         CALL  "#FC_CONTROL_HEATER"
         ( TtA      := "IOC2PLC".TT600,
           TtB      := "IOC2PLC".TT670,
           TtC      := "IOC2PLC".TT680,
           TtD      := "IOC2PLC".TT690,
           TtE      := #Unused_TT,
           TtF      := #Unused_TT,
           Nb_Tt    := 4,
           TS       := #TS,
           ExtCmd   := #ExtCmd,
           cmdEpics := "Epics_to_PLC"."EH60_67-69",
           EH       := "voie 5 chaufferette BV",
           sEpics   := "PLC_to_Epics"."EH60_67-69",
           Object   := "#DATA_HEATERS"."EH60_67-69"
         );
END_REGION

REGION Network 7 (STL): EH97-98 - VB channel 6
   // Dewar, Electrical Heater
         L     2;
         T     "#DATA_HEATERS"."EH97-98".P_TS_Ton;
         T     "#DATA_HEATERS"."EH97-98".P_Pilot_Ton;
         L     5;
         T     "#DATA_HEATERS"."EH97-98".P_TS_Toff;

         SET;
         A     "IOC2PLC".TT970_VALID;
         A     "IOC2PLC".TT980_VALID;
         A     "EPICS_COMM_OK";
         =     #TS;
   // Force the heater ON when the temperature data is not valid
   // (TS = FALSE). The heater will be turned on for 30 s and TS
   // will be forced TRUE for 30 s. This will hopefully raise the
   // temperature enough for Pt100 to be in range (>73 K)
         SET;
         AN    #TS;
         A(;
         A     "#DATA_HEATERS"."EH97-98".XH;
         A     "#DATA_HEATERS"."EH97-98".X;
         O;
         AN    "#DATA_HEATERS"."EH97-98".XH;
         A     "#DATA_HEATERS"."EH97-98".H;
         );
         =     #ExtCmdTrig;
         CALL  TP , "IEC_Timer_EH97-98_DB"
         ( IN := #ExtCmdTrig,
           PT := T#30s,
           Q  := #ExtCmd,
           ET := #tmp_et
         );
         A     #ExtCmd;
         S     #TS;

         CALL  "#FC_CONTROL_HEATER"
         ( TtA      := "IOC2PLC".TT970,
           TtB      := "IOC2PLC".TT980,
           TtC      := #Unused_TT,
           TtD      := #Unused_TT,
           TtE      := #Unused_TT,
           TtF      := #Unused_TT,
           Nb_Tt    := 2,
           TS       := #TS,
           ExtCmd   := #ExtCmd,
           cmdEpics := "Epics_to_PLC"."EH97-98",
           EH       := "voie 6 chaufferette BV",
           sEpics   := "PLC_to_Epics"."EH97-98",
           Object   := "#DATA_HEATERS"."EH97-98"
         );
END_REGION

REGION Network 8 (STL): EH01 - CM channel 1
         L     2;
         T     "#DATA_HEATERS".EH01.P_TS_Ton;
         T     "#DATA_HEATERS".EH01.P_Pilot_Ton;
         L     5;
         T     "#DATA_HEATERS".EH01.P_TS_Toff;

         SET;
         A     "IOC2PLC".TT04_VALID;
         A     "IOC2PLC".TT06_VALID;
         A     "EPICS_COMM_OK";
         =     #TS;

         CALL  "#FC_CONTROL_HEATER"
         ( TtA      := "IOC2PLC".TT04,
           TtB      := "IOC2PLC".TT06,
           TtC      := #Unused_TT,
           TtD      := #Unused_TT,
           TtE      := #Unused_TT,
           TtF      := #Unused_TT,
           Nb_Tt    := 2,
           TS       := #TS,
           ExtCmd   := #ExtCmd,
           cmdEpics := "Epics_to_PLC".EH01,
           EH       := "voie 1 chaufferette CM",
           sEpics   := "PLC_to_Epics".EH01,
           Object   := "#DATA_HEATERS".EH01
         );
END_REGION

REGION Network 9 (STL): EH02 - CM channel 2
         L     2;
         T     "#DATA_HEATERS".EH02.P_TS_Ton;
         T     "#DATA_HEATERS".EH02.P_Pilot_Ton;
         L     5;
         T     "#DATA_HEATERS".EH02.P_TS_Toff;

         SET;
         A     "IOC2PLC".TT05_VALID;
         A     "IOC2PLC".TT07_VALID;
         A     "EPICS_COMM_OK";
         =     #TS;

         CALL  "#FC_CONTROL_HEATER"
         ( TtA      := "IOC2PLC".TT05,
           TtB      := "IOC2PLC".TT07,
           TtC      := #Unused_TT,
           TtD      := #Unused_TT,
           TtE      := #Unused_TT,
           TtF      := #Unused_TT,
           Nb_Tt    := 2,
           TS       := #TS,
           ExtCmd   := #ExtCmd,
           cmdEpics := "Epics_to_PLC".EH02,
           EH       := "voie 2 chaufferette CM",
           sEpics   := "PLC_to_Epics".EH02,
           Object   := "#DATA_HEATERS".EH02
         );
END_REGION

REGION Network 10 (STL): EH10 - CM channel 3
         L     2;
         T     "#DATA_HEATERS".EH10.P_TS_Ton;
         T     "#DATA_HEATERS".EH10.P_Pilot_Ton;
         L     5;
         T     "#DATA_HEATERS".EH10.P_TS_Toff;

         SET;
         A     "IOC2PLC"."CTS:TT10_VALID";
         A     "IOC2PLC"."CTS:TT11_VALID";
         A     "EPICS_COMM_OK";
         =     #TS;

         CALL  "#FC_CONTROL_HEATER"
         ( TtA      := "IOC2PLC"."CTS:TT10",
           TtB      := "IOC2PLC"."CTS:TT11",
           TtC      := #Unused_TT,
           TtD      := #Unused_TT,
           TtE      := #Unused_TT,
           TtF      := #Unused_TT,
           Nb_Tt    := 2,
           TS       := #TS,
           ExtCmd   := #ExtCmd,
           cmdEpics := "Epics_to_PLC".EH10,
           EH       := "voie 3 chaufferette CM",
           sEpics   := "PLC_to_Epics".EH10,
           Object   := "#DATA_HEATERS".EH10
         );
END_REGION

REGION Network 11 (STL): EH20 - CM channel 4
         L     2;
         T     "#DATA_HEATERS".EH20.P_TS_Ton;
         T     "#DATA_HEATERS".EH20.P_Pilot_Ton;
         L     5;
         T     "#DATA_HEATERS".EH20.P_TS_Toff;

         SET;
         A     "IOC2PLC"."CTS:TT20_VALID";
         A     "IOC2PLC"."CTS:TT21_VALID";
         A     "EPICS_COMM_OK";
         =     #TS;

         CALL  "#FC_CONTROL_HEATER"
         ( TtA      := "IOC2PLC"."CTS:TT20",
           TtB      := "IOC2PLC"."CTS:TT21",
           TtC      := #Unused_TT,
           TtD      := #Unused_TT,
           TtE      := #Unused_TT,
           TtF      := #Unused_TT,
           Nb_Tt    := 2,
           TS       := #TS,
           ExtCmd   := #ExtCmd,
           cmdEpics := "Epics_to_PLC".EH20,
           EH       := "voie 4 chaufferette CM",
           sEpics   := "PLC_to_Epics".EH20,
           Object   := "#DATA_HEATERS".EH20
         );
END_REGION

REGION Network 12 (STL): EH918 - CM channel 9
   // Dewar, Electrical Heater
         L     2;
         T     "#DATA_HEATERS"."spare-CM-9".P_TS_Ton;
         T     "#DATA_HEATERS"."spare-CM-9".P_Pilot_Ton;
         L     5;
         T     "#DATA_HEATERS"."spare-CM-9".P_TS_Toff;

         SET;
         A     "IOC2PLC"."CTS:TT20_VALID";
         A     "EPICS_COMM_OK";
         =     #TS;
   // Force the heater ON when the temperature data is not valid
   // (TS = FALSE). The heater will be turned on for 30 s and TS
   // will be forced TRUE for 30 s. This will hopefully raise the
   // temperature enough for Pt100 to be in range (>73 K)
         SET;
         AN    #TS;
         A(;
         A     "#DATA_HEATERS"."spare-CM-9".XH;
         A     "#DATA_HEATERS"."spare-CM-9".X;
         O;
         AN    "#DATA_HEATERS"."spare-CM-9".XH;
         A     "#DATA_HEATERS"."spare-CM-9".H;
         );
         =     #ExtCmdTrig;
         CALL  TP , "IEC_Timer_EH918_DB"
         ( IN := #ExtCmdTrig,
           PT := T#30s,
           Q  := #ExtCmd,
           ET := #tmp_et
         );
         A     #ExtCmd;
         S     #TS;

   _191: CALL  "#FC_CONTROL_HEATER"
         ( TtA      := "IOC2PLC"."CTS:TT20",
           TtB      := #Unused_TT,
           TtC      := #Unused_TT,
           TtD      := #Unused_TT,
           TtE      := #Unused_TT,
           TtF      := #Unused_TT,
           Nb_Tt    := 1,
           TS       := #TS,
           ExtCmd   := #ExtCmd,
           cmdEpics := "Epics_to_PLC"."spare-CM-9",
           EH       := "voie 9 chaufferette CM",
           sEpics   := "PLC_to_Epics"."spare-CM-9",
           Object   := "#DATA_HEATERS"."spare-CM-9"
         );
END_REGION

REGION Network 13 (STL): EH904 - CM channel 11
   // Dewar, Electrical Heater
         L     2;
         T     "#DATA_HEATERS"."spare-CM-11".P_TS_Ton;
         T     "#DATA_HEATERS"."spare-CM-11".P_Pilot_Ton;
         L     5;
         T     "#DATA_HEATERS"."spare-CM-11".P_TS_Toff;

         SET;
         A     "IOC2PLC"."CTS:TT21_VALID";
         A     "EPICS_COMM_OK";
         =     #TS;

   // Force the heater ON when the temperature data is not valid
   // (TS = FALSE). The heater will be turned on for 30 s and TS
   // will be forced TRUE for 30 s. This will hopefully raise the
   // temperature enough for Pt100 to be in range (>73 K)
         SET;
         AN    #TS;
         A(;
         A     "#DATA_HEATERS"."spare-CM-11".XH;
         A     "#DATA_HEATERS"."spare-CM-11".X;
         O;
         AN    "#DATA_HEATERS"."spare-CM-11".XH;
         A     "#DATA_HEATERS"."spare-CM-11".H;
         );
         =     #ExtCmdTrig;
         CALL  TP , "IEC_Timer_EH904_DB"
         ( IN := #ExtCmdTrig,
           PT := T#30s,
           Q  := #ExtCmd,
           ET := #tmp_et
         );
         A     #ExtCmd;
         S     #TS;

         CALL  "#FC_CONTROL_HEATER"
         ( TtA      := "IOC2PLC"."CTS:TT21",
           TtB      := #Unused_TT,
           TtC      := #Unused_TT,
           TtD      := #Unused_TT,
           TtE      := #Unused_TT,
           TtF      := #Unused_TT,
           Nb_Tt    := 1,
           TS       := #TS,
           ExtCmd   := #ExtCmd,
           cmdEpics := "Epics_to_PLC"."spare-CM-11",
           EH       := "voie 11 chaufferette CM",
           sEpics   := "PLC_to_Epics"."spare-CM-11",
           Object   := "#DATA_HEATERS"."spare-CM-11"
         );
END_REGION

REGION Network 14 (STL): EH12 - Coupler 1 flange
   // Dewar, Electrical Heater
         L     2;
         T     "#DATA_HEATERS".EH12.P_TS_Ton;
         T     "#DATA_HEATERS".EH12.P_Pilot_Ton;
         L     5;
         T     "#DATA_HEATERS".EH12.P_TS_Toff;

         L     "PLC_to_Epics".TT120.Visu;
         L     0;
         ==I;
         =     #Enable;
         CALL  "#FC_CONTROL_HEATER"
         ( TtA      := "PLC_to_Epics".TT120.Level,
           TtB      := #Unused_TT,
           TtC      := #Unused_TT,
           TtD      := #Unused_TT,
           TtE      := #Unused_TT,
           TtF      := #Unused_TT,
           Nb_Tt    := 1,
           TS       := #Enable,
           ExtCmd   := #ExtCmd,
           cmdEpics := "Epics_to_PLC".EH12,
           EH       := "EH12 Cpl1",
           sEpics   := "PLC_to_Epics".EH12,
           Object   := "#DATA_HEATERS".EH12
         );
END_REGION

REGION Network 15 (STL): EH22 - Coupler 2 flange
   // Dewar, Electrical Heater
         L     2;
         T     "#DATA_HEATERS".EH22.P_TS_Ton;
         T     "#DATA_HEATERS".EH22.P_Pilot_Ton;
         L     5;
         T     "#DATA_HEATERS".EH22.P_TS_Toff;

         L     "PLC_to_Epics".TT220.Visu;
         L     0;
         ==I;
         =     #Enable;
         CALL  "#FC_CONTROL_HEATER"
         ( TtA      := "PLC_to_Epics".TT220.Level,
           TtB      := #Unused_TT,
           TtC      := #Unused_TT,
           TtD      := #Unused_TT,
           TtE      := #Unused_TT,
           TtF      := #Unused_TT,
           Nb_Tt    := 1,
           TS       := #Enable,
           ExtCmd   := #ExtCmd,
           cmdEpics := "Epics_to_PLC".EH22,
           EH       := "EH22 Cpl2",
           sEpics   := "PLC_to_Epics".EH22,
           Object   := "#DATA_HEATERS".EH22
         );
END_REGION
END_FUNCTION

FUNCTION "Manage_HEATERS" : Void   // FC513, LAD
TITLE = Manage the heaters
{ S7_Optimized_Access := 'FALSE' }
AUTHOR : KG
VERSION : 0.1
BEGIN

REGION Network 1: EH12 & EH22 - Coupler flange cavity 1 and 2
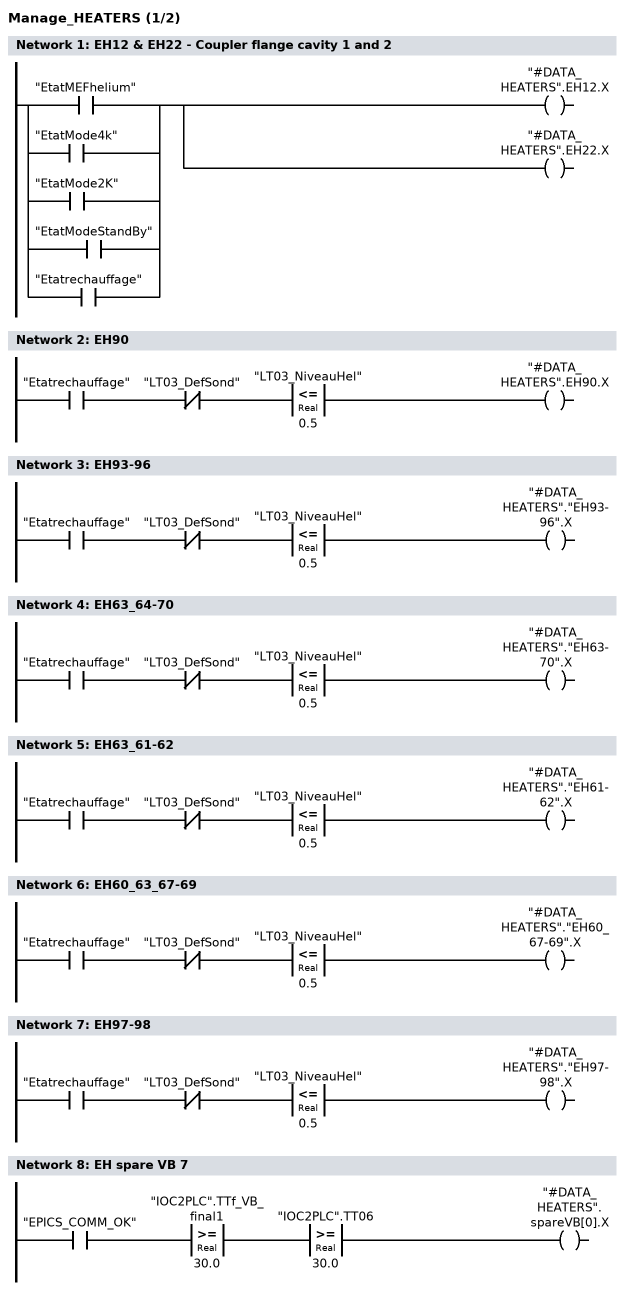
   RUNG wire#powerrail
      Contact( "EtatMEFhelium" )
      wire#w1
      Coil( "#DATA_HEATERS".EH12.X )
   END_RUNG
   RUNG wire#powerrail
      Contact( "EtatMode4k" )
   END_RUNG wire#w1
   RUNG wire#powerrail
      Contact( "EtatMode2K" )
   END_RUNG wire#w1
   RUNG wire#powerrail
      Contact( "EtatModeStandBy" )
   END_RUNG wire#w1
   RUNG wire#powerrail
      Contact( "Etatrechauffage" )
   END_RUNG wire#w1
   RUNG wire#w1
      Coil( "#DATA_HEATERS".EH22.X )
   END_RUNG
   // the same network as SCL:
   "#DATA_HEATERS".EH12.X := "EtatMEFhelium" OR "EtatMode4k" OR "EtatMode2K" OR "EtatModeStandBy" OR "Etatrechauffage";
   "#DATA_HEATERS".EH22.X := "#DATA_HEATERS".EH12.X;
END_REGION

REGION Network 2: EH90
   RUNG wire#powerrail
      Contact( "Etatrechauffage" )
      I_Contact( "LT03_DefSond" )
      { S7_Templates := "SrcType := Real" } LE_Contact(in1 := "LT03_NiveauHel", in2 := 0.5)
      Coil( "#DATA_HEATERS".EH90.X )
   END_RUNG
   // the same network as SCL:
   "#DATA_HEATERS".EH90.X := "Etatrechauffage" AND NOT "LT03_DefSond" AND ("LT03_NiveauHel" <= 0.5);
END_REGION

REGION Network 3: EH93-96
   RUNG wire#powerrail
      Contact( "Etatrechauffage" )
      I_Contact( "LT03_DefSond" )
      { S7_Templates := "SrcType := Real" } LE_Contact(in1 := "LT03_NiveauHel", in2 := 0.5)
      Coil( "#DATA_HEATERS"."EH93-96".X )
   END_RUNG
   // the same network as SCL:
   "#DATA_HEATERS"."EH93-96".X := "Etatrechauffage" AND NOT "LT03_DefSond" AND ("LT03_NiveauHel" <= 0.5);
END_REGION

REGION Network 4: EH63_64-70
   RUNG wire#powerrail
      Contact( "Etatrechauffage" )
      I_Contact( "LT03_DefSond" )
      { S7_Templates := "SrcType := Real" } LE_Contact(in1 := "LT03_NiveauHel", in2 := 0.5)
      Coil( "#DATA_HEATERS"."EH63-70".X )
   END_RUNG
   // the same network as SCL:
   "#DATA_HEATERS"."EH63-70".X := "Etatrechauffage" AND NOT "LT03_DefSond" AND ("LT03_NiveauHel" <= 0.5);
END_REGION

REGION Network 5: EH63_61-62
   RUNG wire#powerrail
      Contact( "Etatrechauffage" )
      I_Contact( "LT03_DefSond" )
      { S7_Templates := "SrcType := Real" } LE_Contact(in1 := "LT03_NiveauHel", in2 := 0.5)
      Coil( "#DATA_HEATERS"."EH61-62".X )
   END_RUNG
   // the same network as SCL:
   "#DATA_HEATERS"."EH61-62".X := "Etatrechauffage" AND NOT "LT03_DefSond" AND ("LT03_NiveauHel" <= 0.5);
END_REGION

REGION Network 6: EH60_63_67-69
   RUNG wire#powerrail
      Contact( "Etatrechauffage" )
      I_Contact( "LT03_DefSond" )
      { S7_Templates := "SrcType := Real" } LE_Contact(in1 := "LT03_NiveauHel", in2 := 0.5)
      Coil( "#DATA_HEATERS"."EH60_67-69".X )
   END_RUNG
   // the same network as SCL:
   "#DATA_HEATERS"."EH60_67-69".X := "Etatrechauffage" AND NOT "LT03_DefSond" AND ("LT03_NiveauHel" <= 0.5);
END_REGION

REGION Network 7: EH97-98
   RUNG wire#powerrail
      Contact( "Etatrechauffage" )
      I_Contact( "LT03_DefSond" )
      { S7_Templates := "SrcType := Real" } LE_Contact(in1 := "LT03_NiveauHel", in2 := 0.5)
      Coil( "#DATA_HEATERS"."EH97-98".X )
   END_RUNG
   // the same network as SCL:
   "#DATA_HEATERS"."EH97-98".X := "Etatrechauffage" AND NOT "LT03_DefSond" AND ("LT03_NiveauHel" <= 0.5);
END_REGION

REGION Network 8: EH spare VB 7
   RUNG wire#powerrail
      Contact( "EPICS_COMM_OK" )
      { S7_Templates := "SrcType := Real" } GE_Contact(in1 := "IOC2PLC".TTf_VB_final1, in2 := 30.0)
      { S7_Templates := "SrcType := Real" } GE_Contact(in1 := "IOC2PLC".TT06, in2 := 30.0)
      Coil( "#DATA_HEATERS".spareVB[0].X )
   END_RUNG
   // the same network as SCL:
   "#DATA_HEATERS".spareVB[0].X := "EPICS_COMM_OK" AND ("IOC2PLC".TTf_VB_final1 >= 30.0) AND ("IOC2PLC".TT06 >= 30.0);
END_REGION

REGION Network 9: EH spare CM 11
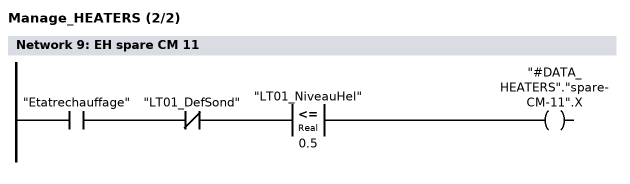
   RUNG wire#powerrail
      Contact( "Etatrechauffage" )
      I_Contact( "LT01_DefSond" )
      { S7_Templates := "SrcType := Real" } LE_Contact(in1 := "LT01_NiveauHel", in2 := 0.5)
      Coil( "#DATA_HEATERS"."spare-CM-11".X )
   END_RUNG
   // the same network as SCL:
   "#DATA_HEATERS"."spare-CM-11".X := "Etatrechauffage" AND NOT "LT01_DefSond" AND ("LT01_NiveauHel" <= 0.5);
END_REGION
END_FUNCTION

FUNCTION "Manage_VALVES" : Void   // FC556, LAD
TITLE = Manage the valves
{ S7_Optimized_Access := 'FALSE' }
AUTHOR : KG
VERSION : 0.1
BEGIN

REGION Network 1: RV90
   // Open the release valve when the pressure is over the threshold
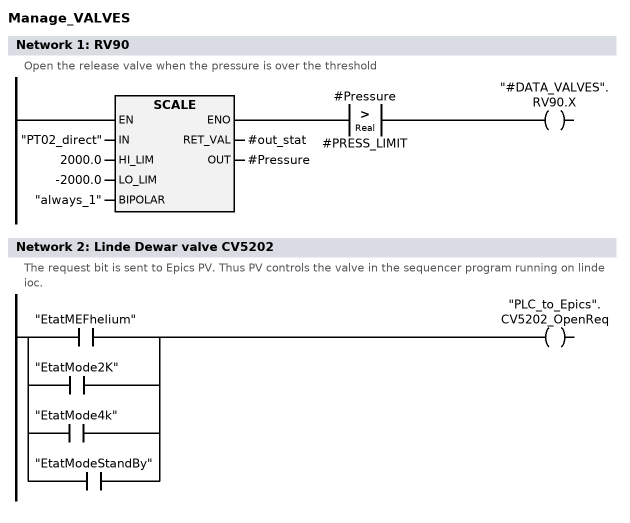
   // ENO of a box is taken as its EN; it also drops when the box reports an error
   #out_stat := SCALE(IN := "PT02_direct",
                      HI_LIM := 2000.0,
                      LO_LIM := -2000.0,
                      BIPOLAR := "always_1",
                      OUT => #Pressure);
   "#DATA_VALVES".RV90.X := #Pressure > #PRESS_LIMIT;
END_REGION

REGION Network 2: Linde Dewar valve CV5202
   // The request bit is sent to Epics PV. Thus PV controls the valve in the sequencer program running on linde ioc.
   RUNG wire#powerrail
      Contact( "EtatMEFhelium" )
      wire#w1
      Coil( "PLC_to_Epics".CV5202_OpenReq )
   END_RUNG
   RUNG wire#powerrail
      Contact( "EtatMode2K" )
   END_RUNG wire#w1
   RUNG wire#powerrail
      Contact( "EtatMode4k" )
   END_RUNG wire#w1
   RUNG wire#powerrail
      Contact( "EtatModeStandBy" )
   END_RUNG wire#w1
   // the same network as SCL:
   "PLC_to_Epics".CV5202_OpenReq := "EtatMEFhelium" OR "EtatMode2K" OR "EtatMode4k" OR "EtatModeStandBy";
END_REGION
END_FUNCTION

ORGANIZATION_BLOCK "Main"   // OB1, STL
TITLE = "Main Program Sweep (Cycle)"
{ S7_Optimized_Access := 'FALSE' }
VERSION : 0.1
BEGIN

REGION Network 1: Set-up the timing pulse for FC_TIMER
         A     "point1sec";
         AN    "point1secMem";
         =     "point1secPls";
         A     "point1sec";
         =     "point1secMem";

         SET;
         A     "oneSec";
         AN    "oneSecMem";
         =     "oneSecPls";
         A     "oneSec";
         =     "oneSecMem";
END_REGION

REGION Network 2: Get data and commands from Epics IOC
         CALL  "Recv_from_Epics";
         NOP   0;
END_REGION

REGION Network 3
         A     "Graph/manuelle";
         JNB   Label_0;
         CALL  "commande vanne";
   Label_0:NOP   0;
END_REGION

REGION Network 4
         CALL  "NIveau Helium&Pression&vide";
         NOP   0;
END_REGION

REGION Network 5
         CALL  "ACQ_CABTF";
         NOP   0;
END_REGION

REGION Network 6
         AN    "Graph/manuelle";
         JNB   Label_1;
         CALL  "grafcet";
   Label_1:NOP   0;
END_REGION

REGION Network 7
         CALL  "Send_to_Epics";
         NOP   0;
END_REGION

REGION Network 8: Instantiate the heaters control
         CALL  "INST_CONTROL_HEATER";
END_REGION

REGION Network 9: Instantiate the valve control
         CALL  "INST_VALVES";
END_REGION

REGION Network 10: Manage the heaters
         CALL  "Manage_HEATERS";
END_REGION

REGION Network 11: Manage the valves
         CALL  "Manage_VALVES";
END_REGION

REGION Network 12
         CALL  "UpdateData2HNOSS";
END_REGION

REGION Network 13: Appeler le bloc de diagnostic système / Call system diagnostics block
         CALL  "RSE_FB", "RSE_DB";
END_REGION

REGION Network 14: Clear INIT flag after the first cycle
         SET;
         R     "INIT";
END_REGION
END_ORGANIZATION_BLOCK

ORGANIZATION_BLOCK "CYC_INT2"   // OB32, LAD
TITLE = Cyclic_1s / "Cyclic Interrupt"
{ S7_Optimized_Access := 'FALSE' }
AUTHOR : KG
VERSION : 0.1
// Call the PID functionswith 1s interval
   VAR_TEMP   // added for the SCL form of the ladder/FBD networks
      _w1 : Bool;
   END_VAR
BEGIN

REGION Network 1: PID regulator for the LN2 screen cooling (CV60)
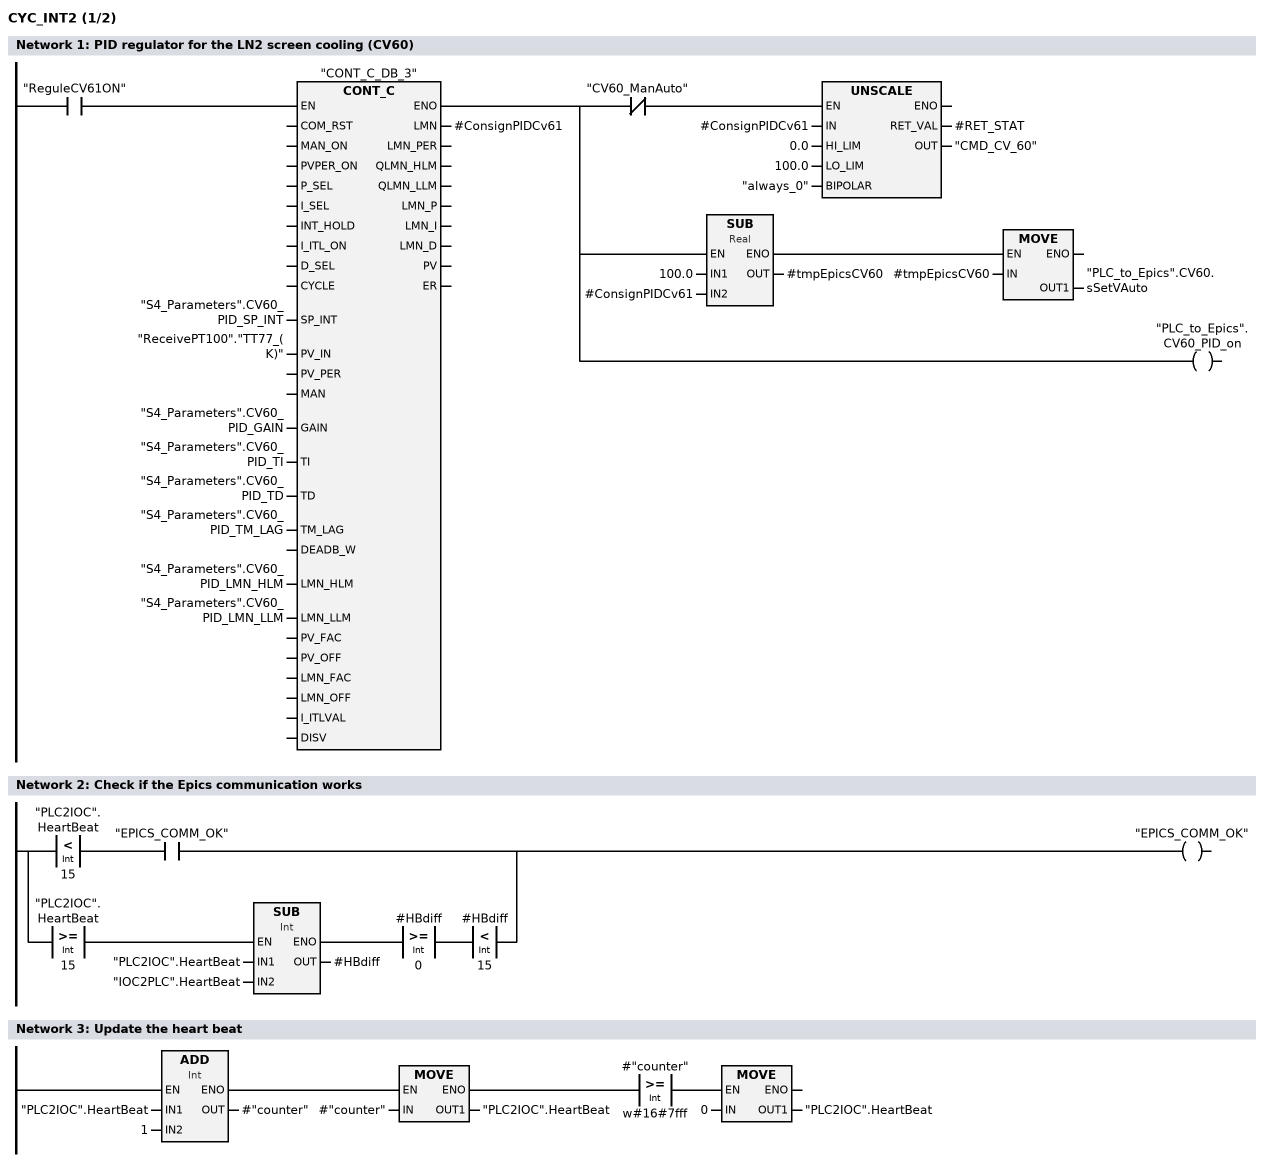
   // ENO of a box is taken as its EN; it also drops when the box reports an error
   #_w1 := "ReguleCV61ON";
   IF #_w1 THEN
       "CONT_C_DB_3"(SP_INT := "S4_Parameters".CV60_PID_SP_INT,   // CONT_C
                     PV_IN := "ReceivePT100"."TT77_(K)",
                     GAIN := "S4_Parameters".CV60_PID_GAIN,
                     TI := "S4_Parameters".CV60_PID_TI,
                     TD := "S4_Parameters".CV60_PID_TD,
                     TM_LAG := "S4_Parameters".CV60_PID_TM_LAG,
                     LMN_HLM := "S4_Parameters".CV60_PID_LMN_HLM,
                     LMN_LLM := "S4_Parameters".CV60_PID_LMN_LLM,
                     LMN => #ConsignPIDCv61);
   END_IF;
   IF #_w1 AND NOT "CV60_ManAuto" THEN
       #RET_STAT := UNSCALE(IN := #ConsignPIDCv61,
                            HI_LIM := 0.0,
                            LO_LIM := 100.0,
                            BIPOLAR := "always_0",
                            OUT => "CMD_CV_60");
   END_IF;
   IF #_w1 THEN
       #tmpEpicsCV60 := 100.0 - #ConsignPIDCv61;
       "PLC_to_Epics".CV60.sSetVAuto := #tmpEpicsCV60;
   END_IF;
   "PLC_to_Epics".CV60_PID_on := #_w1;
END_REGION

REGION Network 2: Check if the Epics communication works
   // ENO of a box is taken as its EN; it also drops when the box reports an error
   #_w1 := "PLC2IOC".HeartBeat >= 15;
   IF #_w1 THEN #HBdiff := "PLC2IOC".HeartBeat - "IOC2PLC".HeartBeat; END_IF;
   "EPICS_COMM_OK" := (#_w1 AND (#HBdiff >= 0) AND (#HBdiff < 15)) OR (("PLC2IOC".HeartBeat < 15) AND "EPICS_COMM_OK");
END_REGION

REGION Network 3: Update the heart beat
   RUNG wire#powerrail
      { S7_Templates := "SrcType := Int"; S7_GenerateENO := "TRUE" } Add(in1 := "PLC2IOC".HeartBeat, in2 := 1, out => #"counter")
      { S7_GenerateENO := "TRUE" } Move(in := #"counter", out1 => "PLC2IOC".HeartBeat)
      { S7_Templates := "SrcType := Int" } GE_Contact(in1 := #"counter", in2 := w#16#7fff)
      { S7_GenerateENO := "TRUE" } Move(in := 0, out1 => "PLC2IOC".HeartBeat)
   END_RUNG
   // the same network as SCL:
   // ENO of a box is taken as its EN; it also drops when the box reports an error
   #"counter" := "PLC2IOC".HeartBeat + 1;
   "PLC2IOC".HeartBeat := #"counter";
   IF #"counter" >= w#16#7fff THEN "PLC2IOC".HeartBeat := 0; END_IF;
END_REGION

REGION Network 4: Check if the communicationto HNOSS PLC works
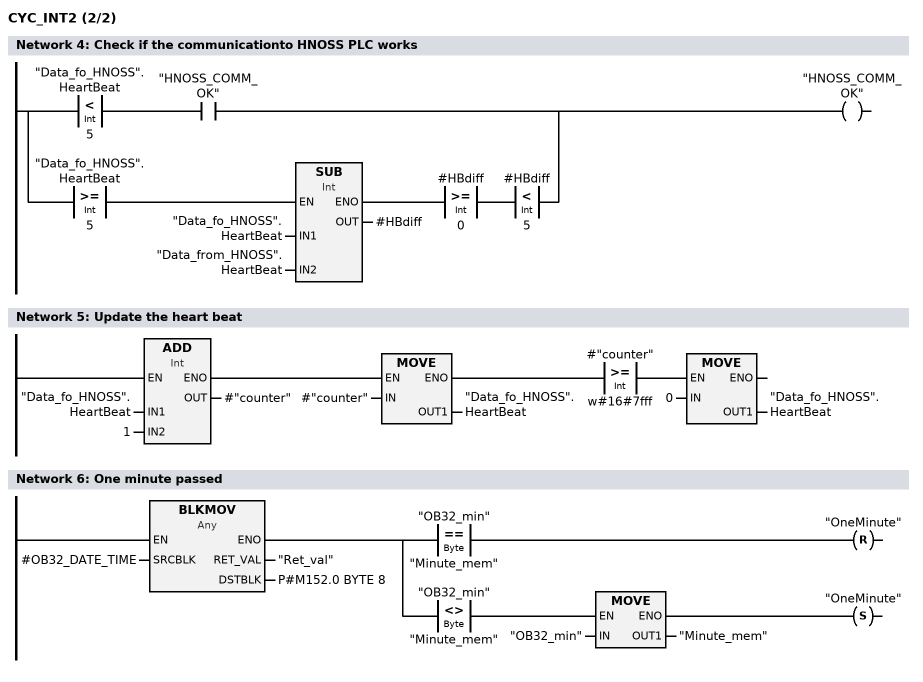
   // ENO of a box is taken as its EN; it also drops when the box reports an error
   #_w1 := "Data_fo_HNOSS".HeartBeat >= 5;
   IF #_w1 THEN #HBdiff := "Data_fo_HNOSS".HeartBeat - "Data_from_HNOSS".HeartBeat; END_IF;
   "HNOSS_COMM_OK" := (#_w1 AND (#HBdiff >= 0) AND (#HBdiff < 5)) OR (("Data_fo_HNOSS".HeartBeat < 5) AND "HNOSS_COMM_OK");
END_REGION

REGION Network 5: Update the heart beat
   RUNG wire#powerrail
      { S7_Templates := "SrcType := Int"; S7_GenerateENO := "TRUE" } Add(in1 := "Data_fo_HNOSS".HeartBeat, in2 := 1, out => #"counter")
      { S7_GenerateENO := "TRUE" } Move(in := #"counter", out1 => "Data_fo_HNOSS".HeartBeat)
      { S7_Templates := "SrcType := Int" } GE_Contact(in1 := #"counter", in2 := w#16#7fff)
      { S7_GenerateENO := "TRUE" } Move(in := 0, out1 => "Data_fo_HNOSS".HeartBeat)
   END_RUNG
   // the same network as SCL:
   // ENO of a box is taken as its EN; it also drops when the box reports an error
   #"counter" := "Data_fo_HNOSS".HeartBeat + 1;
   "Data_fo_HNOSS".HeartBeat := #"counter";
   IF #"counter" >= w#16#7fff THEN "Data_fo_HNOSS".HeartBeat := 0; END_IF;
END_REGION

REGION Network 6: One minute passed
   // ENO of a box is taken as its EN; it also drops when the box reports an error
   "Ret_val" := BLKMOV(SRCBLK := #OB32_DATE_TIME, DSTBLK => P#M152.0 BYTE 8);
   IF "OB32_min" = "Minute_mem" THEN "OneMinute" := FALSE; END_IF;
   #_w1 := "OB32_min" <> "Minute_mem";
   IF #_w1 THEN
       "Minute_mem" := "OB32_min";
       "OneMinute" := TRUE;
   END_IF;
END_REGION
END_ORGANIZATION_BLOCK

ORGANIZATION_BLOCK "CYC_INT5"   // OB35, LAD
TITLE = "Cyclic Interrupt"
{ S7_Optimized_Access := 'FALSE' }
VERSION : 0.1
// Period 100 ms
   VAR_TEMP   // added for the SCL form of the ladder/FBD networks
      _w1 : Bool;
      _w2 : Bool;
   END_VAR
BEGIN

REGION Network 1
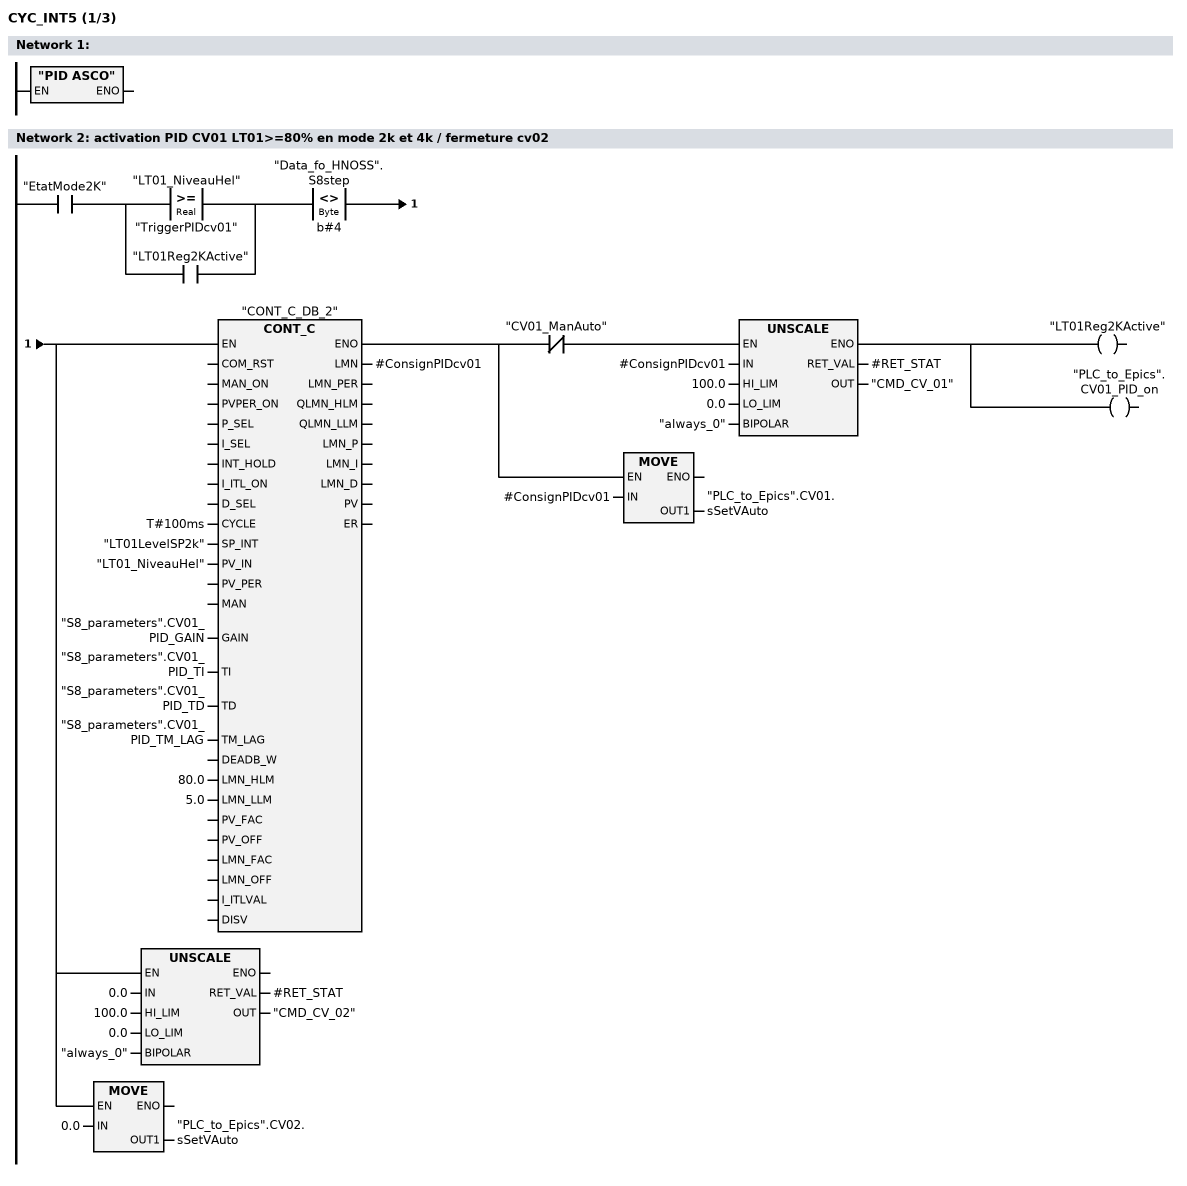
   RUNG wire#powerrail
      "PID ASCO"()
   END_RUNG
   // the same network as SCL:
   "PID ASCO"();
END_REGION

REGION Network 2: activation PID CV01 LT01>=80% en mode 2k et 4k / fermeture cv02
   // ENO of a box is taken as its EN; it also drops when the box reports an error
   #_w1 := "EtatMode2K" AND (("LT01_NiveauHel" >= "TriggerPIDcv01") OR "LT01Reg2KActive") AND ("Data_fo_HNOSS".S8step <> b#4);
   IF #_w1 THEN
       "CONT_C_DB_2"(CYCLE := T#100ms,   // CONT_C
                     SP_INT := "LT01LevelSP2k",
                     PV_IN := "LT01_NiveauHel",
                     GAIN := "S8_parameters".CV01_PID_GAIN,
                     TI := "S8_parameters".CV01_PID_TI,
                     TD := "S8_parameters".CV01_PID_TD,
                     TM_LAG := "S8_parameters".CV01_PID_TM_LAG,
                     LMN_HLM := 80.0,
                     LMN_LLM := 5.0,
                     LMN => #ConsignPIDcv01);
   END_IF;
   #_w2 := #_w1 AND NOT "CV01_ManAuto";
   IF #_w2 THEN
       #RET_STAT := UNSCALE(IN := #ConsignPIDcv01,
                            HI_LIM := 100.0,
                            LO_LIM := 0.0,
                            BIPOLAR := "always_0",
                            OUT => "CMD_CV_01");
   END_IF;
   "LT01Reg2KActive" := #_w2;
   "PLC_to_Epics".CV01_PID_on := #_w2;
   IF #_w1 THEN
       "PLC_to_Epics".CV01.sSetVAuto := #ConsignPIDcv01;
       #RET_STAT := UNSCALE(IN := 0.0, HI_LIM := 100.0, LO_LIM := 0.0, BIPOLAR := "always_0", OUT => "CMD_CV_02");
       "PLC_to_Epics".CV02.sSetVAuto := 0.0;
   END_IF;
END_REGION

REGION Network 3: activation PID CV03 LT03>=80%
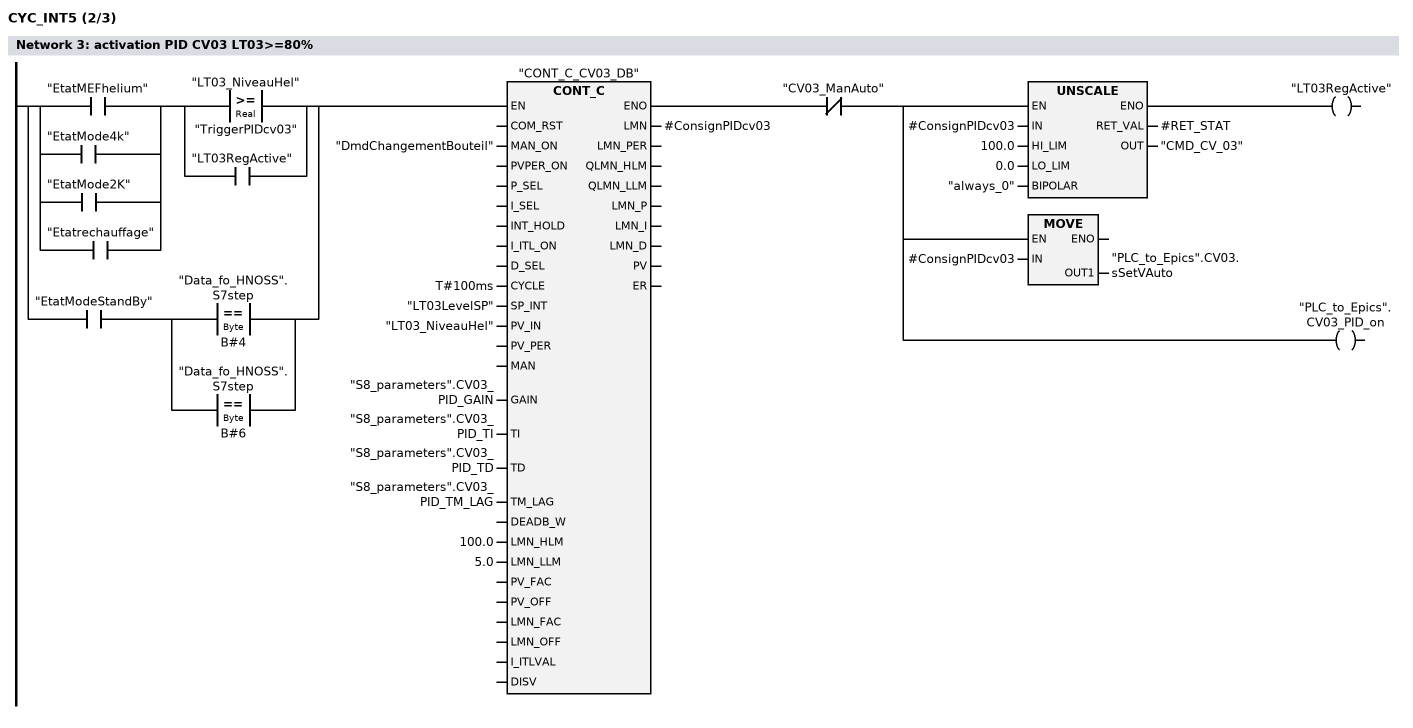
   // ENO of a box is taken as its EN; it also drops when the box reports an error
   #_w1 := (("EtatMEFhelium" OR "EtatMode4k" OR "EtatMode2K" OR "Etatrechauffage") AND (("LT03_NiveauHel" >= "TriggerPIDcv03") OR "LT03RegActive")) OR ("EtatModeStandBy" AND (("Data_fo_HNOSS".S7step = B#4) OR ("Data_fo_HNOSS".S7step = B#6)));
   IF #_w1 THEN
       "CONT_C_CV03_DB"(MAN_ON := "DmdChangementBouteil",   // CONT_C
                        CYCLE := T#100ms,
                        SP_INT := "LT03LevelSP",
                        PV_IN := "LT03_NiveauHel",
                        GAIN := "S8_parameters".CV03_PID_GAIN,
                        TI := "S8_parameters".CV03_PID_TI,
                        TD := "S8_parameters".CV03_PID_TD,
                        TM_LAG := "S8_parameters".CV03_PID_TM_LAG,
                        LMN_HLM := 100.0,
                        LMN_LLM := 5.0,
                        LMN => #ConsignPIDcv03);
   END_IF;
   #_w2 := #_w1 AND NOT "CV03_ManAuto";
   IF #_w2 THEN
       #RET_STAT := UNSCALE(IN := #ConsignPIDcv03,
                            HI_LIM := 100.0,
                            LO_LIM := 0.0,
                            BIPOLAR := "always_0",
                            OUT => "CMD_CV_03");
   END_IF;
   "LT03RegActive" := #_w2;
   IF #_w2 THEN "PLC_to_Epics".CV03.sSetVAuto := #ConsignPIDcv03; END_IF;
   "PLC_to_Epics".CV03_PID_on := #_w2;
END_REGION

REGION Network 4: activation PID CV02 LT01>=80%
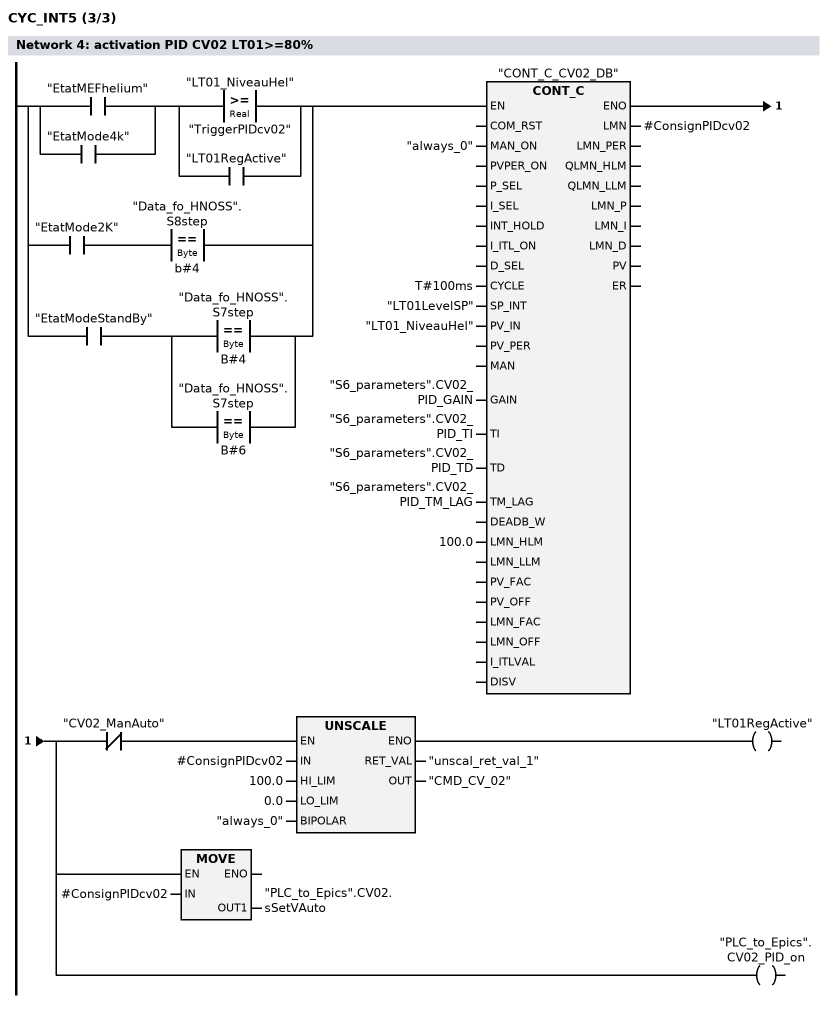
   // ENO of a box is taken as its EN; it also drops when the box reports an error
   #_w1 := (("EtatMEFhelium" OR "EtatMode4k") AND (("LT01_NiveauHel" >= "TriggerPIDcv02") OR "LT01RegActive")) OR ("EtatMode2K" AND ("Data_fo_HNOSS".S8step = b#4)) OR ("EtatModeStandBy" AND (("Data_fo_HNOSS".S7step = B#4) OR ("Data_fo_HNOSS".S7step = B#6)));
   IF #_w1 THEN
       "CONT_C_CV02_DB"(MAN_ON := "always_0",   // CONT_C
                        CYCLE := T#100ms,
                        SP_INT := "LT01LevelSP",
                        PV_IN := "LT01_NiveauHel",
                        GAIN := "S6_parameters".CV02_PID_GAIN,
                        TI := "S6_parameters".CV02_PID_TI,
                        TD := "S6_parameters".CV02_PID_TD,
                        TM_LAG := "S6_parameters".CV02_PID_TM_LAG,
                        LMN_HLM := 100.0,
                        LMN => #ConsignPIDcv02);
   END_IF;
   #_w2 := #_w1 AND NOT "CV02_ManAuto";
   IF #_w2 THEN
       "unscal_ret_val_1" := UNSCALE(IN := #ConsignPIDcv02,
                               HI_LIM := 100.0,
                               LO_LIM := 0.0,
                               BIPOLAR := "always_0",
                               OUT => "CMD_CV_02");
   END_IF;
   "LT01RegActive" := #_w2;
   IF #_w1 THEN "PLC_to_Epics".CV02.sSetVAuto := #ConsignPIDcv02; END_IF;
   "PLC_to_Epics".CV02_PID_on := #_w1;
END_REGION
END_ORGANIZATION_BLOCK

ORGANIZATION_BLOCK "HW_INT0"   // OB40, LAD
TITLE = "Hardware Interrupt"
{ S7_Optimized_Access := 'FALSE' }
VERSION : 0.1
BEGIN
END_ORGANIZATION_BLOCK

ORGANIZATION_BLOCK "I/O_FLT1"   // OB82, LAD
TITLE = "I/O Point Fault"
{ S7_Optimized_Access := 'FALSE' }
VERSION : 0.1
BEGIN

REGION Network 1 (STL): Appeler le bloc de diagnostic système / Call system diagnostics block
         CALL  "RSE_FB", "RSE_DB";
END_REGION
END_ORGANIZATION_BLOCK

ORGANIZATION_BLOCK "OBNL_FLT"   // OB85, LAD
TITLE = "Organization Block (OB) Not Loaded Fault"
{ S7_Optimized_Access := 'FALSE' }
VERSION : 0.1
BEGIN
END_ORGANIZATION_BLOCK

ORGANIZATION_BLOCK "RACK_FLT"   // OB86, LAD
TITLE = "Loss Of Rack Fault"
{ S7_Optimized_Access := 'FALSE' }
VERSION : 0.1
BEGIN

REGION Network 1 (STL): Appeler le bloc de diagnostic système / Call system diagnostics block
         CALL  "RSE_FB", "RSE_DB";
END_REGION
END_ORGANIZATION_BLOCK

ORGANIZATION_BLOCK "COMPLETE RESTART"   // OB100, STL
TITLE = "Complete Restart"
{ S7_Optimized_Access := 'FALSE' }
VERSION : 0.1
BEGIN

REGION Network 1
         SET;
         S     "INIT";
END_REGION

REGION Network 2: S5 parameters
         L     "Epics_to_PLC".S5_P_FT552_MIN_GB.cSetV;
         T     "PLC_to_Epics".S5_P_FT552_MIN_GB.sSetV;
         L     "Epics_to_PLC".S5_P_FT552_MIN_C.cSetV;
         T     "PLC_to_Epics".S5_P_FT552_MIN_C.sSetV;
         L     "Epics_to_PLC".S5_P_FT552_MAX_GB.cSetV;
         T     "PLC_to_Epics".S5_P_FT552_MAX_GB.sSetV;
         L     "Epics_to_PLC".S5_P_FT552_MAX_C.cSetV;
         T     "PLC_to_Epics".S5_P_FT552_MAX_C.sSetV;
END_REGION

REGION Network 3: PID settings
         L     "Epics_to_PLC".TrigPID_CV01.cSetV;
         T     "TriggerPIDcv01";
         L     "Epics_to_PLC".TrigPID_CV02.cSetV;
         T     "TriggerPIDcv02";
         L     "Epics_to_PLC".TrigPID_CV03.cSetV;
         T     "TriggerPIDcv03";
         L     "Epics_to_PLC".PID_LT01_CV01_SP.cSetV;
         T     "LT01LevelSP2k";
         L     "Epics_to_PLC".PID_LT03_CV03_SP.cSetV;
         T     "LT03LevelSP";
         L     "Epics_to_PLC".PID_LT01_CV02_SP.cSetV;
         T     "LT01LevelSP";
         L     "Epics_to_PLC".PID_PT01_CV550_SP.cSetV;
         T     "RéguleASCO02_SP";
         T     "Data_fo_HNOSS".SP_PT01_MKS2;
END_REGION

REGION Network 4: CV550
         L     "Epics_to_PLC".CV550.cSetv;
         T     "PLC_to_Epics".CV550.sSetV;
         T     "Data_fo_HNOSS".CV550_MKS2;
END_REGION

REGION Network 5: S8 parameters
         L     "Epics_to_PLC".S8_P_CV01.cSetV;
         T     "PLC_to_Epics".S8_P_CV01.sSetV;
END_REGION
END_ORGANIZATION_BLOCK

(* ===== HMI "HMI_RT_1" =====

graphic list "Vanne horizontale maxi_0": 1 'Vanne horizontale verte_2'; 0 'Vanne horizontale rouge_2'; 2 'Vanne horizontale rouge_2'; 3 'Vanne horizontale verte_2'; 4 'Vanne horizontale grise_2'; 5 'Vanne horizontale grise_2'

ScreenModuleEditorView "Bloc Vanne horizontale" 1024x768
   GraphicIOField "Modèle_Champ E/S graphique_13" at 10,10 size 50x35
*)

(* ===== HMI "HMI_RT_1" =====

graphic list "Vanne verticale maxi_0": 1 'Vanne verticale verte_1'; 2 'Vanne verticale rouge_1'; 0 'Vanne verticale rouge_1'; 3 'Vanne verticale verte_1'; 4 'Vanne verticale grise_1'; 5 'Vanne verticale grise_1'

ScreenModuleEditorView "Bloc Vanne verticale" 1024x768
   GraphicIOField "Champ E/S graphique_10" at 10,10 size 35x50
*)